REGION Network 4: Time handle
   // Es werden die Absolutwerte der Zeiten berechnet um sie dann vergleichen zu 
   // können. Intervallzeiten sind minimal 10sec. Sonst Störung "Zeitwert falsch"!
   // Bei Spaltfiltern max Laufzeit 20sec.,Min Pausenzeit 300sec.und kein Dauerbetrieb
   // möglich!
   //-----
         SET;
         R     #Temp_WrongTimevalue;
   //-----
         L     #IN_Values.RunTime;
         T     #Temp_RunTime;
         L     #IN_Values.PauseTime;
         T     #Temp_PauseTime;
   //-----
   // Absolutwerte berechnen
   //-----
         CALL  T_CONV
         ( IN  := #Temp_RunTime,
           OUT := #Temp_Runtime_ms
         );
   //-----
         CALL  T_CONV
         ( IN  := #Temp_PauseTime,
           OUT := #Temp_Pausetime_ms
         );
   //-----
         SET;
         R     #Temp_IO_Status.No_Pausetime;
   //-----
         O(;
         L     #Temp_Runtime_ms;
         L     0;
         ==I;
         );
         O(;
         L     #Temp_Pausetime_ms;
         L     0;
         ==I;
         );
         S     #Temp_IO_Status.No_Pausetime;
   //-----
   // Zeiten limitieren
   //-----
         L     #Temp_Runtime_ms;
         L     10000;  // 10 sec
         <D;
         S     #Temp_WrongTimevalue;  // Antrieb STOP!!!
         JCN   RTime;
   //-----
         L     S5T#10S;
         T     #Temp_RunTime;
   //-----
   RTime:NOP   0;
   //-----
         L     #Temp_Pausetime_ms;
         L     10000;  // 10.0 sec
         <D;
         S     #Temp_WrongTimevalue;  // Antrieb STOP!!!
   //-----
         JCN   PTime;
         L     S5T#10S;
         T     #Temp_PauseTime;
   //-----
   PTime:NOP   0;
   //-----
         O     #Temp_IO_Status.No_Pausetime;
         R     #Temp_WrongTimevalue;
   //-----
         A     #Temp_WrongTimevalue;
         AN    #Temp_IO_Fault.FLT_wrong_Timevalue;
         S     #Temp_IO_Fault.FLT_wrong_Timevalue;
         S     #IO_NewFault;
END_REGION

REGION Network 5
   //-----
         O     #Temp_IO_Fault.FLT_Motorprotection;
         O     #Temp_IO_Fault.FLT_FrequencyConverter;
         O     #Temp_IO_Fault.FLT_MaxLTripTray;
         O     #Temp_IO_Fault.FLT_wrong_Timevalue;
         =     #Temp_IO_Status.FaultLevel_3;
   //-----
END_REGION

REGION Network 6: Error handling
   //-----
         O     #Temp_IO_Fault.FLT_Motorprotection;
         O     #Temp_IO_Fault.FLT_FrequencyConverter;
         O     #Temp_IO_Fault.FLT_MaxLTripTray;
         O     #Temp_IO_Fault.FLT_wrong_Timevalue;
         O     #Temp_IO_Fault.Mes_Min_Level;
         =     #Temp_IO_Status.FLT_Exist;
   //-----
         O     #Temp_IO_Fault.FLT_Motorprotection;
         O     #Temp_IO_Fault.FLT_FrequencyConverter;
         O     #Temp_IO_Fault.FLT_MaxLTripTray;
         O     #Temp_IO_Fault.FLT_wrong_Timevalue;
         O     #Temp_IO_Fault.Mes_Min_Level;
         S     #Temp_IO_Status.Reset_Intervall;
         S     #IO_FaultLevel_3;
   //-----
END_REGION

REGION Network 7: Desicion intervall or not!
   //-----
         O(;
         A     #IN_Request_Filling;
         A     #IN_Values.Config_bit_Filling_ON;
         AN    #IN_Values.Config_bit_Filling_Int;
         );
   //-----
         O(;
         A     #IN_Request_Feed;
         A     #IN_Values.Config_bit_Charging_ON;
         AN    #IN_Values.Config_bit_Charging_Int;
         );
   //-----
         O(;
         A     #IN_Request_Cooling;
         A     #IN_Values.Config_bit_Cooling_ON;
         AN    #IN_Values.Config_bit_Cooling_Int;
         );
   //-----
         O(;
         A     #IN_Request_Heating;
         A     #IN_Values.Config_bit_Heating_ON;
         AN    #IN_Values.config_bit_Heating_Int;
         );
   //-----
         O     #Temp_IO_Status.No_Pausetime;
         S     #Temp_IO_Status.Reset_Intervall;
   //-----
END_REGION

REGION Network 8: Reset Intervall / Angefordert setzen
   //-----
         ON    #Temp_ReleaseDrive;
         ON    #IN_Release;
         O     #Temp_IO_Status.Reset_Intervall;
         R     #Temp_IO_Status.Run;
         R     #Temp_IO_Status.Pause;
         R     #Temp_IO_Status.Reset_Intervall;
   //-----
END_REGION

REGION Network 9: Wiedereinschaltsperre
   //-----
         ON    #IN_ControlVoltage;
         FP    #Temp_IO_Status.Ramp_CVoltage_Off;
         S     #Temp_IO_Status.Start_Startupdelay;
         R     #Temp_IO_Status.Disable_Start;
         R     #IN_TimerDrive;
   //-----
         ON    #IN_Values.Config_bit_Converter;
         O     #IN_TimerDrive;
         A     #Temp_IO_Status.Start_Startupdelay;
         R     #Temp_IO_Status.Disable_Start;
         R     #Temp_IO_Status.Start_Startupdelay;
   //-----
         A     #Temp_IO_Status.Start_Startupdelay;
         JCN   Lauf;
   //-----
         A     #Temp_IO_Status.Disable_Start;
         L     S5T#10S;
         SD    #IN_TimerDrive;
   //-----
         SET;
         S     #Temp_IO_Status.Disable_Start;
   //-----
         A     #IN_TimerDrive;
         A     #Temp_IO_Status.Start_Startupdelay;
         R     #Temp_IO_Status.Start_Startupdelay;
         R     #Temp_IO_Status.Disable_Start;
   //-----
END_REGION

REGION Network 10: Laufzeit
   //-----
   Lauf: NOP   0;
   //-----
         A     #Temp_ReleaseDrive;
         AN    #Temp_IO_Status.Pause;
         AN    #Temp_IO_Status.Start_Startupdelay;
         JCN   Paus;
   //-----
         A     #Temp_IO_Status.Run;
         L     #Temp_RunTime;
         SD    #IN_TimerDrive;
   //-----
         SET;
         S     #Temp_IO_Status.Run;
   //-----
         A     #IN_TimerDrive;
         JCN   Ausg;
   //-----
         SET;
         R     #Temp_IO_Status.Run;
         R     #IN_TimerDrive;
   //-----
END_REGION

REGION Network 11: Pause
   //-----
   Paus: NOP   0;
   //-----
         A     #Temp_ReleaseDrive;
         AN    #Temp_IO_Status.Run;
         AN    #Temp_IO_Status.Start_Startupdelay;
         JCN   Ausg;
   //-----
         A     #Temp_IO_Status.Pause;
         L     #Temp_PauseTime;
         SD    #IN_TimerDrive;
   //-----
         SET;
         S     #Temp_IO_Status.Pause;
   //-----
         A     #IN_TimerDrive;
         JCN   Ausg;
   //-----
         SET;
         R     #Temp_IO_Status.Pause;
         R     #IN_TimerDrive;
   //-----
END_REGION

REGION Network 12: Output mainscontactor
   //-----
   Ausg: NOP   0;
   //-----
         O(;  // generel switch ON without frequency converter
         O     #Temp_IO_Status.No_Pausetime;
         O     #Temp_IO_Status.Run;
         A     #Temp_ReleaseDrive;
         AN    #Temp_IO_Fault.Mes_Min_Level;
         AN    #Temp_IO_Fault.FLT_wrong_Timevalue;
         AN    #Temp_IO_Fault.FLT_MaxLTripTray;
         AN    #IN_Values.Config_bit_Converter;
         );
   //-----
         O(;  // generel switch ON withfrequency converter
         A     #IN_ControlVoltage;
         AN    #Temp_IO_Status.Start_Startupdelay;
         A     #IN_Values.Config_bit_Converter;
         );
         AN    #Temp_IO_Fault.FLT_Motorprotection;
   //-----
         =     #Temp_Out_MainsContactor;
         =     #OUT_MainsContactor;
   //-----
END_REGION

REGION Network 13: Ouput release frequency converter
   //-----
         O     #Temp_IO_Status.No_Pausetime;
         O     #Temp_IO_Status.Run;
         A     #Temp_ReleaseDrive;
         A     #Temp_Out_MainsContactor;
         A     #IN_Values.Config_bit_Converter;
         AN    #Temp_IO_Fault.Mes_Min_Level;
         AN    #Temp_IO_Fault.FLT_wrong_Timevalue;
         AN    #Temp_IO_Fault.FLT_MaxLTripTray;
         AN    #Temp_IO_Fault.FLT_FrequencyConverter;
         A     #IN_FaultFreqConverter;
         =     #OUT_Release_FConverter;
         =     #Temp_Release_FConverter;
   //-----
END_REGION

REGION Network 14: State of drive: 1-> ON; 2-> Faulty; 3->Selected but not ON
   //-----
         AN    #IN_Values.Config_bit_Converter;
         A     #Temp_Out_MainsContactor;
         O     #Temp_Release_FConverter;
         L     1;
         JC    tran;
   //-----
         O     #Temp_IO_Status.FLT_Exist;
         L     2;
         JC    tran;
   //-----
         AN(;
         AN    #IN_Values.Config_bit_Converter;
         A     #Temp_Out_MainsContactor;
         O     #Temp_Release_FConverter;
         );
         AN    #Temp_IO_Status.FLT_Exist;
         A     #Temp_IO_Status.Switch_Drive_ON_OFF;
         L     3;
         JC    tran;
   //-----
         L     0;
   //-----
   tran: T     #Temp_IO_Status.State_Drive;
   //-----
END_REGION

REGION Network 15: Save data
   //-----
         CALL  BLKMOV
         ( SRCBLK  := #Temp_IO_Status,
           RET_VAL := #ERROR_CODE,
           DSTBLK  := #Anyzeiger1
         );
   //-----
         CALL  BLKMOV
         ( SRCBLK  := #Temp_IO_Fault,
           RET_VAL := #ERROR_CODE,
           DSTBLK  := #Anyzeiger2
         );
   //-----
END_REGION
END_FUNCTION

FUNCTION "FC122_EdgeFilter" : Void   // FC122, STL
TITLE = Control of several auxiliary drives of a pouring machine
{ S7_Optimized_Access := 'FALSE' }
AUTHOR : KT242
FAMILY : RS_KK
NAME : Drive
VERSION : 1.5
   VAR_INPUT
      IN_Release : Bool;   // Genarelly release 0f the drive (Operation mode)
      IN_Reset_fault : Bool;   // Signal to quit fault within function block
      IN_Fault_Motorprotection : Bool;   // Input fault motorprotection of drive
      IN_DifPressure : Bool;   // Input fault difference pressure
      IN_TimerDrive : Timer;   // Timer of general timing of the drive
      Values : "UDT710_EdgeFilter";
   END_VAR
   VAR_OUTPUT
      OUT_MainsContactor : Bool;   // Ouput mainscontactor drive or frequency converter
   END_VAR
   VAR_IN_OUT
      IO_Status : ANY;   // Stores the state of the drive
      IO_NewFault : Bool;
      IO_FaultLevel_3 : Bool;
      IO_Faults : ANY;
   END_VAR
   VAR_TEMP
      Temp_IO_Status : "UDT100_EdgeFilter";
      ERROR_CODE : Int;   // Error state of systemfunction "BLKMOV" Blockmove
      Anyzeiger1 : ANY;   // Pointer to copy thr array "IO_Status" and "Temp_IO_Status"
      Anyzeiger2 : ANY;   // Pointer to copy thr array "IO_Status" and "Temp_IO_Status"
      Temp_IO_Fault : "UDT1801_EdgeFilter";
      Temp_RunTime : S5Time;   // Flag runtime drive
      Temp_PauseTime : S5Time;   // Flag pause time
      Temp_Runtime_ms : Time;   // Flag runtime drive in millisecond
      Temp_Pausetime_ms : Time;   // Flag pause time drive in millisecond
      Temp_ReleaseDrive : Bool;   // Flag release activation drive
      Temp_Fault_Drive : Bool;
      Temp_MainsContactor : Bool;
   END_VAR
BEGIN

REGION Network 1: Saved data integration
   // Änderungen:
   // -------------------------------------------------------------------------------
   // Bei der Verwendung der Umwälzpumpe als Speisepumpe wurde dieses bei Min. 
   // Füllstand ausgeshaltet, auch wenn dies im Zyklus auftrat. Hierdurch wurden dann 
   // auch die Materialpumpen abgeschaltet.
   // v.d.Geest     25.02.2003
   // -------------------------------------------------------------------------------
   // Bei einer Ansteuerung mit Frequenzumrichter wurde nicht auf die 
   // Störungsauswertung des Umrichters gewartet bevor die Freigabe gegeben wurde. 
   // Hierdurch kam es zu Störungen bei jedem einschalten des Aggregates.
   // A. Jäger      21.11.2003
   //-----
         LAR1;
         L;
         LAR2;
   //-----
         L     W[AR2, P#0.0];  // Bytes
         T     W[AR1, P#0.0];
         L     W[AR2, P#2.0];  // Amount of bytes
         T     W[AR1, P#2.0];
         L     W[AR2, P#4.0];  // Block no,
         T     W[AR1, P#4.0];
         L     D[AR2, P#6.0];  // Startadress of datas
         T     D[AR1, P#6.0];
   //-----
         CALL  BLKMOV
         ( SRCBLK  := #Anyzeiger1,
           RET_VAL := #ERROR_CODE,
           DSTBLK  := #Temp_IO_Status
         );
   //-----
         LAR1;
         L;
         LAR2;
   //-----
         L     W[AR2, P#0.0];  // Bytes
         T     W[AR1, P#0.0];
         L     W[AR2, P#2.0];  // Amount of bytes
         T     W[AR1, P#2.0];
         L     W[AR2, P#4.0];  // Block no,
         T     W[AR1, P#4.0];
         L     D[AR2, P#6.0];  // Startadress of datas
         T     D[AR1, P#6.0];
   //-----
         CALL  BLKMOV
         ( SRCBLK  := #Anyzeiger2,
           RET_VAL := #ERROR_CODE,
           DSTBLK  := #Temp_IO_Fault
         );
   //-----
END_REGION

REGION Network 2: Fault motorprotection
   //-----
         AN    #Values.Config_Exist;
         R     #Temp_IO_Fault.FLT_Motorprotection;
         R     #Temp_IO_Fault.FLT_MaxPressureDiff;
         R     #Temp_IO_Fault.FLT_wrong_Timevalue;
         R     #Temp_IO_Status.FLT_Exist;
         R     #Temp_IO_Status.Pause;
         R     #Temp_IO_Status.Run;
         JC    Ausg;
   //-----
END_REGION

REGION Network 3: Release drive
   //-----
         O     #Temp_IO_Status.Switch_Drive_ON_OFF;
         A     #IN_Release;
         =     #Temp_ReleaseDrive;
   //-----
END_REGION

REGION Network 4: Faults
   //-----
         A     #IN_Reset_fault;
         R     #Temp_IO_Fault.FLT_Motorprotection;
         R     #Temp_IO_Fault.FLT_MaxPressureDiff;
         R     #Temp_IO_Fault.FLT_wrong_Timevalue;
   //-----
         A     #IN_Fault_Motorprotection;
         AN    #Temp_IO_Fault.FLT_Motorprotection;
         S     #Temp_IO_Fault.FLT_Motorprotection;
         S     #Temp_IO_Status.Reset_Intervall;
         S     #IO_NewFault;
   //-----
         AN    #IN_DifPressure;
         A     #Values.Config_DifPress;
         A     #Temp_ReleaseDrive;
         AN    #Temp_IO_Fault.FLT_MaxPressureDiff;
         S     #Temp_IO_Fault.FLT_MaxPressureDiff;
         S     #Temp_IO_Status.Reset_Intervall;
         S     #IO_NewFault;
   //-----
END_REGION

REGION Network 5
   //-----
         O     #Temp_IO_Fault.FLT_Motorprotection;
         O     #Temp_IO_Fault.FLT_MaxPressureDiff;
         O     #Temp_IO_Fault.FLT_wrong_Timevalue;
         =     #Temp_IO_Status.FLT_Exist;
         =     #Temp_Fault_Drive;
         =     #Temp_IO_Status.FaultLevel_3;
         S     #IO_FaultLevel_3;
   //-----
END_REGION

REGION Network 6: Time handle
   // Es werden die Absolutwerte der Zeiten berechnet um sie dann vergleichen zu 
   // können. Intervallzeiten sind minimal 10sec. Sonst Störung "Zeitwert falsch"!
   // Bei Spaltfiltern max Laufzeit 20sec.,Min Pausenzeit 300sec.und kein Dauerbetrieb
   // möglich!
   //-----
         SET;
         R     #Temp_IO_Fault.FLT_wrong_Timevalue;
   //-----
         L     #Values.RunTime;
         T     #Temp_RunTime;
         L     #Values.PauseTime;
         T     #Temp_PauseTime;
   //-----
   // Absolutwerte berechnen
   //-----
         CALL  T_CONV
         ( IN  := #Temp_RunTime,
           OUT := #Temp_Runtime_ms
         );
   //-----
         CALL  T_CONV
         ( IN  := #Temp_PauseTime,
           OUT := #Temp_Pausetime_ms
         );
   //-----
   // Zeiten limitieren
   //-----
         L     #Temp_Runtime_ms;
         L     20000;  // 20.0 sec
         >D;
         S     #Temp_IO_Fault.FLT_wrong_Timevalue;  // Antrieb STOP!!!
   //-----
         JCN   RTimeS;
         L     S5T#20S;
         T     #Temp_RunTime;
   RTimeS:NOP   0;
   //-----
         L     #Temp_Pausetime_ms;
         L     L#300000;  // 300.0 sec
         <D;
         S     #Temp_IO_Fault.FLT_wrong_Timevalue;  // Antrieb STOP!!!
   //-----
         JCN   PTimeS;
         L     S5T#5M;
         T     #Temp_PauseTime;
   //-----
   PTimeS:NOP   0;
   //-----
END_REGION

REGION Network 7: Reset Intervall / Angefordert setzen
   //-----
         ON    #Temp_ReleaseDrive;
         O     #Temp_IO_Status.Reset_Intervall;
         R     #Temp_IO_Status.Run;
         R     #Temp_IO_Status.Pause;
         R     #Temp_IO_Status.Reset_Intervall;
   //-----
END_REGION

REGION Network 8: Laufzeit
   Lauf: NOP   0;
         A     #Temp_ReleaseDrive;
         AN    #Temp_IO_Status.Pause;
         JCN   Paus;
   //
         A     #Temp_IO_Status.Run;
         L     #Temp_RunTime;
         SD    #IN_TimerDrive;
   //
         SET;
         S     #Temp_IO_Status.Run;
   //
         A     #IN_TimerDrive;
         JCN   Ausg;
         SET;
         R     #Temp_IO_Status.Run;
         R     #IN_TimerDrive;
END_REGION

REGION Network 9: Pause
   Paus: NOP   0;
         A     #Temp_ReleaseDrive;
         AN    #Temp_IO_Status.Run;
         JCN   Ausg;
   //
         A     #Temp_IO_Status.Pause;
         L     #Temp_PauseTime;
         SD    #IN_TimerDrive;
   //
         SET;
         S     #Temp_IO_Status.Pause;
   //
         A     #IN_TimerDrive;
         JCN   Ausg;
         SET;
         R     #Temp_IO_Status.Pause;
         R     #IN_TimerDrive;
END_REGION

REGION Network 10: Output mainscontactor
   Ausg: NOP   0;
   //
         A     #Temp_IO_Status.Run;  // generell Eingeschaltet ohne FU
         A     #Temp_IO_Status.Switch_Drive_ON_OFF;
         A     #IN_Release;
         AN    #Temp_IO_Fault.FLT_wrong_Timevalue;
         AN    #Temp_IO_Fault.FLT_MaxPressureDiff;
         AN    #Temp_IO_Fault.FLT_Motorprotection;
         A     #Values.Config_Exist;
         =     #OUT_MainsContactor;
         =     #Temp_MainsContactor;
END_REGION

REGION Network 11: State of drive: 1-> ON; 2->Faulty; 3->Selected but not on
   //-----
         A     #Temp_MainsContactor;
         L     1;
         JC    tran;
   //-----
         A     #Temp_Fault_Drive;
         L     2;
         JC    tran;
   //-----
         A     #Temp_IO_Status.Switch_Drive_ON_OFF;
         L     3;
         JC    tran;
   //-----
         L     0;
   //-----
   tran: T     #Temp_IO_Status.State_Drive;
END_REGION

REGION Network 12: Save data
         CALL  BLKMOV
         ( SRCBLK  := #Temp_IO_Status,
           RET_VAL := #ERROR_CODE,
           DSTBLK  := #Anyzeiger1
         );
   //
         CALL  BLKMOV
         ( SRCBLK  := #Temp_IO_Fault,
           RET_VAL := #ERROR_CODE,
           DSTBLK  := #Anyzeiger2
         );
   //
END_REGION
END_FUNCTION

FUNCTION "FC123_FeedingPump" : Void   // FC123, STL
TITLE = Control of several auxiliary drives of a pouring machine
{ S7_Optimized_Access := 'FALSE' }
AUTHOR : KT242
FAMILY : RS_KK
NAME : Drive
VERSION : 1.5
   VAR_INPUT
      IN_Release : Bool;   // Genarelly release 0f the drive (Operation mode)
      IN_ControlVoltage : Bool;   // Signal delay activation frequency converter (protection after emergency-stop)
      IN_Reset_fault : Bool;   // Signal to quit fault within function block
      IN_ComponentDeselected : Bool;   // is the component deselected? -> Fault Group 1 -> Groupe 3
      IN_Request_Feed : Bool;   // Request switch on drive if componenten pump start up
      IN_Request_Filling : Bool;   // Request switch on drive for filling
      IN_Request_Bypass : Bool;   // Request switch on drive for bypass circulation
      IN_Fault_Motorprotection : Bool;   // Input fault motorprotection of drive
      IN_FaultFreqConverter : Bool;   // Input fault frequency converter of drive
      IN_DryRun : Bool;   // Input fault Min_Level or dry run
      IN_MaxLevelTray : Bool;   // Input fault max. filling level tray
      IN_MaxPressure : Bool;   // Input Max pressure switch
      IN_TempRelease : Bool;   // Input Min. Temperature reacht for switch on
      IN_TimerDrive : Timer;   // Timer of general timing of the drive
      IN_TimerStartUpFConv : Timer;   // Timer of delay start up frequency converter
      Values : "UDT710_FeedingPump";
   END_VAR
   VAR_OUTPUT
      OUT_MainsContactor : Bool;   // Ouput mainscontactor drive or frequency converter
      OUT_Release_FConverter : Bool;   // Output release of frequncy converter to control rotation speed
   END_VAR
   VAR_IN_OUT
      IO_Status : ANY;   // Stores the state of the drive
      IO_NewFault : Bool;
      IO_FaultLevel_1 : Bool;
      IO_FaultLevel_3 : Bool;
      IO_Faults : ANY;
   END_VAR
   VAR_TEMP
      Temp_IO_Status : "UDT100_FeedingPump";
      ERROR_CODE : Int;   // Error state of systemfunction "BLKMOV" Blockmove
      Anyzeiger1 : ANY;   // Pointer to copy thr array "IO_Status" and "Temp_IO_Status"
      Anyzeiger2 : ANY;   // Pointer to copy thr array "IO_Status" and "Temp_IO_Status"
      Temp_IO_Fault : "UDT1801_FeedingPump";
      Temp_RunTime : S5Time;   // Flag runtime drive
      Temp_PauseTime : S5Time;   // Flag pause time
      Temp_Runtime_ms : Time;   // Flag runtime drive in millisecond
      Temp_Pausetime_ms : Time;   // Flag pause time drive in millisecond
      Temp_ReleaseDrive : Bool;   // Flag release activation drive
      Temp_Fault_Drive : Bool;
      Temp_WrongTimevalue : Bool;
      Temp_MainsContactor : Bool;
      Temp_Release_FConverter : Bool;
   END_VAR
BEGIN

REGION Network 1: Saved data integration
   // Änderungen:
   // -------------------------------------------------------------------------------
   // Bei der Verwendung der Umwälzpumpe als Speisepumpe wurde dieses bei Min. 
   // Füllstand ausgeshaltet, auch wenn dies im Zyklus auftrat. Hierdurch wurden dann 
   // auch die Materialpumpen abgeschaltet.
   // v.d.Geest     25.02.2003
   // -------------------------------------------------------------------------------
   // Bei einer Ansteuerung mit Frequenzumrichter wurde nicht auf die 
   // Störungsauswertung des Umrichters gewartet bevor die Freigabe gegeben wurde. 
   // Hierdurch kam es zu Störungen bei jedem einschalten des Aggregates.
   // A. Jäger      21.11.2003
   //-----
         LAR1;
         L;
         LAR2;
   //-----
         L     W[AR2, P#0.0];  // Bytes
         T     W[AR1, P#0.0];
         L     W[AR2, P#2.0];  // Amount of bytes
         T     W[AR1, P#2.0];
         L     W[AR2, P#4.0];  // Block no,
         T     W[AR1, P#4.0];
         L     D[AR2, P#6.0];  // Startadress of datas
         T     D[AR1, P#6.0];
   //-----
         CALL  BLKMOV
         ( SRCBLK  := #Anyzeiger1,
           RET_VAL := #ERROR_CODE,
           DSTBLK  := #Temp_IO_Status
         );
   //-----
         LAR1;
         L;
         LAR2;
   //-----
         L     W[AR2, P#0.0];  // Bytes
         T     W[AR1, P#0.0];
         L     W[AR2, P#2.0];  // Amount of bytes
         T     W[AR1, P#2.0];
         L     W[AR2, P#4.0];  // Block no,
         T     W[AR1, P#4.0];
         L     D[AR2, P#6.0];  // Startadress of datas
         T     D[AR1, P#6.0];
   //-----
         CALL  BLKMOV
         ( SRCBLK  := #Anyzeiger2,
           RET_VAL := #ERROR_CODE,
           DSTBLK  := #Temp_IO_Fault
         );
   //-----
END_REGION

REGION Network 2: Fault motorprotection
   //-----
         AN    #Values.Config_Exist;
         R     #Temp_IO_Fault.FLT_Motorprotection;
         R     #Temp_IO_Fault.FLT_FrequencyConverter;
         R     #Temp_IO_Fault.FLT_MaxLTripTray;
         R     #Temp_IO_Fault.FLT_Dryrunsafety;
         R     #Temp_IO_Fault.FLT_wrong_Timevalue;
         R     #Temp_IO_Fault.FLT_MaxPressure;
         R     #Temp_IO_Fault.Mes_Min_temp;
         R     #Temp_IO_Status.FLT_Exist;
         R     #Temp_IO_Status.Pause;
         R     #Temp_IO_Status.Run;
         JC    Ausg;
   //-----
END_REGION

REGION Network 3: Release drive
   //-----
         O(;
         A     #IN_Request_Filling;
         A     #Values.Config_Filling;
         A     #Temp_IO_Status.Switch_Drive_ON_OFF;
         );
         O(;
         A     #IN_Request_Bypass;
         A     #Values.Config_Bypass;
         A     #Temp_IO_Status.Switch_Drive_ON_OFF;
         );
         O(;
         A     #Temp_IO_Status.Switch_Drive_ON_OFF;
         A     #Values.Config_ManualSwitchON;
         );
         O(;
         A     #IN_Request_Feed;
         );
         A     #IN_Release;
         =     #Temp_ReleaseDrive;
   //-----
END_REGION

REGION Network 4: Faults
   //-----
         A     #IN_Reset_fault;
         R     #Temp_IO_Fault.FLT_Motorprotection;
         R     #Temp_IO_Fault.FLT_FrequencyConverter;
         R     #Temp_IO_Fault.FLT_MaxLTripTray;
         R     #Temp_IO_Fault.FLT_Dryrunsafety;
         R     #Temp_IO_Fault.FLT_wrong_Timevalue;
         R     #Temp_IO_Fault.FLT_MaxPressure;
   //-----
         A     #IN_Fault_Motorprotection;
         AN    #Temp_IO_Fault.FLT_Motorprotection;
         S     #Temp_IO_Fault.FLT_Motorprotection;
         S     #IO_NewFault;
   //-----
         A     #IN_ControlVoltage;
         AN    #Temp_IO_Fault.FLT_wrong_Timevalue;
         AN    #Temp_IO_Status.Start_Startupdelay;
         L     S5T#5S;
         SD    #IN_TimerStartUpFConv;
   //-----
         A     #IN_TimerStartUpFConv;
         AN    #IN_FaultFreqConverter;
         A     #Temp_ReleaseDrive;
         A     #Values.Config_WithFC;
         AN    #Temp_IO_Fault.FLT_FrequencyConverter;
         S     #Temp_IO_Fault.FLT_FrequencyConverter;
         S     #IO_NewFault;
   //-----
         AN    #IN_MaxLevelTray;
         A     #Temp_ReleaseDrive;
         AN    #Temp_IO_Fault.FLT_MaxLTripTray;
         S     #Temp_IO_Fault.FLT_MaxLTripTray;
         S     #IO_NewFault;
   //-----
         AN    #IN_DryRun;
         A     #Temp_ReleaseDrive;
         AN    #Temp_IO_Fault.FLT_Dryrunsafety;
         S     #Temp_IO_Fault.FLT_Dryrunsafety;
         S     #IO_NewFault;
   //-----
         AN    #IN_MaxPressure;
         AN    #Temp_IO_Fault.FLT_MaxPressure;
         S     #Temp_IO_Fault.FLT_MaxPressure;
         S     #IO_NewFault;
   //-----
         AN    #IN_TempRelease;
         A     #Temp_ReleaseDrive;
         AN    #Temp_IO_Fault.Mes_Min_temp;
         S     #Temp_IO_Fault.Mes_Min_temp;
         S     #IO_NewFault;
   //-----
         A     #IN_TempRelease;
         ON    #Temp_ReleaseDrive;
         R     #Temp_IO_Fault.Mes_Min_temp;
   //-----
         A     #Temp_IO_Fault.Mes_Min_temp;
         R     #Temp_ReleaseDrive;
   //-----
END_REGION

REGION Network 5: A fault group 1 exist
   //-----
         O     #Temp_IO_Fault.FLT_MaxLTripTray;
         O     #Temp_IO_Fault.FLT_MaxPressure;
         O     #Temp_IO_Fault.FLT_Dryrunsafety;
         AN    #IN_ComponentDeselected;
         =     #Temp_IO_Status.FaultLevel_1;
   //-----
         O     #Temp_IO_Fault.FLT_MaxLTripTray;
         O     #Temp_IO_Fault.FLT_MaxPressure;
         O     #Temp_IO_Fault.FLT_Dryrunsafety;
         A     #IN_ComponentDeselected;
         O     #Temp_IO_Fault.FLT_Motorprotection;
         O     #Temp_IO_Fault.FLT_FrequencyConverter;
         O     #Temp_IO_Fault.FLT_wrong_Timevalue;
         =     #Temp_IO_Status.FaultLevel_3;
   //-----
END_REGION

REGION Network 6: Time handle
   // Es werden die Absolutwerte der Zeiten berechnet um sie dann vergleichen zu 
   // können. Intervallzeiten sind minimal 10sec. Sonst Störung "Zeitwert falsch"!
   // Bei Spaltfiltern max Laufzeit 20sec.,Min Pausenzeit 300sec.und kein Dauerbetrieb
   // möglich!
   //-----
         SET;
         R     #Temp_WrongTimevalue;
   //-----
         L     #Values.RunTime;
         T     #Temp_RunTime;
         L     #Values.PauseTime;
         T     #Temp_PauseTime;
   //-----
   // Absolutwerte berechnen
   //-----
         CALL  T_CONV
         ( IN  := #Temp_RunTime,
           OUT := #Temp_Runtime_ms
         );
   //-----
         CALL  T_CONV
         ( IN  := #Temp_PauseTime,
           OUT := #Temp_Pausetime_ms
         );
   //-----
         SET;
         R     #Temp_IO_Status.No_Pausetime;
   //-----
         O(;
         L     #Temp_Runtime_ms;
         L     0;
         ==I;
         );
         O(;
         L     #Temp_Pausetime_ms;
         L     0;
         ==I;
         );
         S     #Temp_IO_Status.No_Pausetime;
   //-----
   // Zeiten limitieren
   //-----
         L     #Temp_Runtime_ms;
         L     10000;  // 10 sec
         <D;
         S     #Temp_WrongTimevalue;  // Antrieb STOP!!!
         JCN   nLi1;
   //-----
         L     S5T#10S;
         T     #Temp_RunTime;
   //-----
   nLi1: L     #Temp_Pausetime_ms;
         L     10000;  // 10.0 sec
         <D;
         S     #Temp_WrongTimevalue;  // Antrieb STOP!!!
         JCN   nLi2;
   //-----
         L     S5T#10S;
         T     #Temp_PauseTime;
         JU    nLi2;
   //-----
   nLi2: NOP   0;
   //-----
         AN    #Temp_WrongTimevalue;
         R     #Temp_IO_Fault.FLT_wrong_Timevalue;
   //-----
         A     #Temp_WrongTimevalue;
         AN    #Temp_IO_Status.No_Pausetime;
         AN    #Temp_IO_Fault.FLT_wrong_Timevalue;
         S     #Temp_IO_Fault.FLT_wrong_Timevalue;
         S     #IO_NewFault;
   //-----
END_REGION

REGION Network 7: Error handling
   //-----
         O     #Temp_IO_Fault.FLT_Motorprotection;
         O     #Temp_IO_Fault.FLT_FrequencyConverter;
         O     #Temp_IO_Fault.FLT_MaxLTripTray;
         O     #Temp_IO_Fault.FLT_Dryrunsafety;
         O     #Temp_IO_Fault.FLT_wrong_Timevalue;
         =     #Temp_IO_Status.FLT_Exist;
         =     #Temp_Fault_Drive;
   //-----
         O     #Temp_IO_Fault.FLT_Motorprotection;
         O     #Temp_IO_Fault.FLT_FrequencyConverter;
         O     #Temp_IO_Fault.FLT_Dryrunsafety;
         O     #Temp_IO_Fault.FLT_MaxLTripTray;
         O     #Temp_IO_Fault.FLT_wrong_Timevalue;
         S     #Temp_IO_Status.Reset_Intervall;
         S     #IO_FaultLevel_3;
   //-----
END_REGION

REGION Network 8: Desicion intervall or not!
         O(;
         A     #IN_Request_Filling;
         A     #Values.Config_Filling;
         A     #Temp_IO_Status.Switch_Drive_ON_OFF;
         );
         O     #IN_Request_Feed;
         O     #Temp_IO_Status.No_Pausetime;
         S     #Temp_IO_Status.Reset_Intervall;
END_REGION

REGION Network 9: Reset Intervall / Angefordert setzen
   //-----
         ON    #Temp_ReleaseDrive;
         ON    #IN_Release;
         O     #Temp_IO_Status.Reset_Intervall;
         R     #Temp_IO_Status.Run;
         R     #Temp_IO_Status.Pause;
         R     #Temp_IO_Status.Reset_Intervall;
   //-----
END_REGION

REGION Network 10: Wiedereinschaltsperre
   //-----
         ON    #IN_ControlVoltage;
         FP    #Temp_IO_Status.Ramp_CVoltage_Off;
         S     #Temp_IO_Status.Start_Startupdelay;
         R     #Temp_IO_Status.Disable_Start;
         R     #IN_TimerDrive;
   //-----
         ON    #Values.Config_WithFC;
         O     #IN_TimerDrive;
         A     #Temp_IO_Status.Start_Startupdelay;
         R     #Temp_IO_Status.Disable_Start;
         R     #Temp_IO_Status.Start_Startupdelay;
   //-----
         A     #Temp_IO_Status.Start_Startupdelay;
         JCN   Lauf;
   //-----
         A     #Temp_IO_Status.Disable_Start;
         L     S5T#10S;
         SD    #IN_TimerDrive;
   //-----
         SET;
         S     #Temp_IO_Status.Disable_Start;
   //-----
         A     #IN_TimerDrive;
         A     #Temp_IO_Status.Start_Startupdelay;
         R     #Temp_IO_Status.Start_Startupdelay;
         R     #Temp_IO_Status.Disable_Start;
   //-----
END_REGION

REGION Network 11: Laufzeit
   Lauf: NOP   0;
         A     #Temp_ReleaseDrive;
         AN    #Temp_IO_Status.Pause;
         AN    #Temp_IO_Status.Start_Startupdelay;
         JCN   Paus;
   //
         A     #Temp_IO_Status.Run;
         L     #Temp_RunTime;
         SD    #IN_TimerDrive;
   //
         SET;
         S     #Temp_IO_Status.Run;
   //
         A     #IN_TimerDrive;
         JCN   Ausg;
         SET;
         R     #Temp_IO_Status.Run;
         R     #IN_TimerDrive;
END_REGION

REGION Network 12: Pause
   //-----
   Paus: NOP   0;
   //-----
         A     #Temp_ReleaseDrive;
         AN    #Temp_IO_Status.Run;
         AN    #Temp_IO_Status.Start_Startupdelay;
         JCN   Ausg;
   //-----
         A     #Temp_IO_Status.Pause;
         L     #Temp_PauseTime;
         SD    #IN_TimerDrive;
   //-----
         SET;
         S     #Temp_IO_Status.Pause;
   //-----
         A     #IN_TimerDrive;
         JCN   Ausg;
   //-----
         SET;
         R     #Temp_IO_Status.Pause;
         R     #IN_TimerDrive;
   //-----
END_REGION

REGION Network 13: Output mainscontactor
   //-----
   Ausg: NOP   0;
   //-----
         O(;  // generel switch ON without frequency converter
         O     #Temp_IO_Status.No_Pausetime;
         O     #Temp_IO_Status.Run;
         A     #Temp_ReleaseDrive;
         A(;  // If Filling is aktiv the dryrun must switched
         A     #IN_Request_Filling;
         A     #Values.Config_Filling;
         A     #Temp_IO_Status.Switch_Drive_ON_OFF;
         ON    #Temp_IO_Fault.FLT_Dryrunsafety;
         );
         AN    #Temp_IO_Fault.FLT_wrong_Timevalue;
         AN    #Temp_IO_Fault.FLT_MaxLTripTray;
         AN    #Values.Config_WithFC;
         );
         O(;  // generel switch ON withfrequency converter
         A     #IN_ControlVoltage;
         AN    #Temp_IO_Status.Start_Startupdelay;
         A     #Values.Config_WithFC;
         );
         AN    #Temp_IO_Fault.FLT_Motorprotection;
         A     #Values.Config_Exist;
   //-----
         =     #OUT_MainsContactor;
         =     #Temp_MainsContactor;
   //-----
END_REGION

REGION Network 14: Ouput release frequency converter
   //-----
         O     #Temp_IO_Status.No_Pausetime;
         O     #Temp_IO_Status.Run;
         A     #Temp_ReleaseDrive;
         A     #Temp_MainsContactor;
         A     #Values.Config_WithFC;
         A(;  // If Filling is aktiv the dryrun must switched
         A     #IN_Request_Filling;
         A     #Values.Config_Filling;
         A     #Temp_IO_Status.Switch_Drive_ON_OFF;
         ON    #Temp_IO_Fault.FLT_Dryrunsafety;
         );
         AN    #Temp_IO_Fault.FLT_wrong_Timevalue;
         AN    #Temp_IO_Fault.FLT_MaxLTripTray;
         AN    #Temp_IO_Fault.FLT_FrequencyConverter;
         A     #IN_FaultFreqConverter;
         A     #Values.Config_Exist;
         =     #OUT_Release_FConverter;
         =     #Temp_Release_FConverter;
   //-----
END_REGION

REGION Network 15: State of drive: 1-> ON; 2-> Faulty; 3->Selected but not ON
   //-----
         AN    #Values.Config_WithFC;
         A     #Temp_MainsContactor;
         O     #Temp_Release_FConverter;
         L     1;
         JC    tran;
   //-----
         A     #Temp_Fault_Drive;
         L     2;
         JC    tran;
   //-----
         A     #Temp_IO_Status.Switch_Drive_ON_OFF;
         L     3;
         JC    tran;
   //-----
         L     0;
   //-----
   tran: T     #Temp_IO_Status.State_Drive;
   //-----
END_REGION

REGION Network 16: Save data
   //-----
         CALL  BLKMOV
         ( SRCBLK  := #Temp_IO_Status,
           RET_VAL := #ERROR_CODE,
           DSTBLK  := #Anyzeiger1
         );
   //-----
         CALL  BLKMOV
         ( SRCBLK  := #Temp_IO_Fault,
           RET_VAL := #ERROR_CODE,
           DSTBLK  := #Anyzeiger2
         );
   //-----
END_REGION
END_FUNCTION

FUNCTION "FC126_write_ProCan" : Void   // FC126, STL
TITLE = Write to IO-Interface of ProCan modul
{ S7_Optimized_Access := 'FALSE' }
AUTHOR : KT242
FAMILY : RS_KK
NAME : WRProcan
VERSION : 1.1
   VAR_TEMP
      Nullmerker : Byte;   // Zwischenmerker mit dem Wert "0" zum ablöschen bei gestörter Übertragung
      ERROR_CODE : DInt;   // Störungszustand der Systemfunktion "FILL" Blockmove
      Temp_ToolAdr : Int;
      Temp_PS_offset : Int;
      TempShotWithMaterial_M1 : Bool;
      TempShotWithMaterial_M2 : Bool;
      Temp_OperationMode : Bool;
      ControlBitShot : Byte;
      Temp_MH_OutputSignals : Word;
      TempMH_Bit : DWord;
      Temp_MH_Shot_MH01 : Bool;
      Temp_MH_Shot_MH02 : Bool;
      Temp_MH_Shot_MH03 : Bool;
      Temp_MH_Shot_MH04 : Bool;
      Temp_MH_Shot_MH05 : Bool;
      Temp_MH_Shot_MH06 : Bool;
      Temp_MH_Shot_MH07 : Bool;
      Temp_MH_Shot_MH08 : Bool;
      Temp_MH_Shot_MH09 : Bool;
      Temp_MH_Shot_MH10 : Bool;
      Temp_CorrValue : Real;
      Temp_Error : Bool;
      TempFlowIndex : Byte;
      TemRetBLKMOV : Int;
      TempTandem : Word;
      Dummy : Bool;
      TempNozzelBitCirc : Byte;
      TempNozzelBitShot : Byte;
      TempAdrNozzel : Int;
      TempNozzelBitForce : Byte;
      ControlByteCtrlCP : Byte;
      ThrottleGap : Int;
      TempNozzelBitRelease : Byte;
      ShotTime_M1 : DInt;
      ControlFlowIndex : Byte;
      ControlBitCP : Byte;
      Temp_CycleRunning : Array[1..16] of Bool;
   END_VAR
BEGIN

REGION Network 1: Write data flow 1
   //----------------------------------------------------------------------
   // Check if the communication partner is ready for
   // data transfer to ProCan
   // ---------------------------------------------------------------------
         AN    "PN_FlowRate".Component[1].FlowC_F.Active;
         JC    ed01;
   //-----------------------------------------------------------------
   // Flow set value
   //-----------------------------------------------------------------
         L     0;
         L     "PN_FlowRate".Component[1].FlowC_F.Address;
         <>D;
         JCN   qp01;
         SLD   3;
         LAR1;
         L     0;
         A     "TM_pulse_2PointAdjust_C1";
         JC    _2point_C1;
         L     "DB613_Komponent_State".FlowPump[1];
   _2point_C1:T     PQD [ AR1 , P#0.0 ];

   //---------------------------------------------------------------------
   // Quick pressure build up
   //---------------------------------------------------------------------
   qp01: L     0;
         L     "PN_FlowRate".Component[1].FlowC_F.Address;
         <>D;
         JCN   fi01;
         L     4;
         +D;
         SLD   3;
         LAR1;
         L     "DB613_Komponent_State".FlowPumpQPB[1];
         T     PQD[AR1, P#0.0];

         L     0;
         L     "PN_FlowRate".Component[1].FlowC_F.Address;
         <>D;
         JCN   fi01;
         L     8;
         +D;
         SLD   3;
         LAR1;
         L     "DB613_Komponent_State".PressurePumpQPB[1];
         T     PQD [ AR1 , P#0.0 ];

   //--- Pressure from external device ???
   //    L     0
   //    L     "DB1233_ProCanIO_Flow".AddressFlow[1].Ref_Act_PressureQPB
   //    <I
   //    SPBN  fi01
   //    SLD   3
   //    LAR1
   //    L     DB60.DBW    2
   //    L     10
   //    *D
   //    T     PAW [AR1,P#0.0]

   //-----------------------------------------------------------------
   // Flow-Index: Enableclosedloop; Start quick pressure build up
   //-----------------------------------------------------------------
   fi01: L     0;
         T     #ControlFlowIndex;

   //-----------------------------------------
   // Enableclosedloop
   //-----------------------------------------
         AN    "DB613_Komponent_State".MeteringPump[1].Enableclosedloop;
         JC    SDA1;
         L     2#0000_0010;
         L     #ControlFlowIndex;
         OW;
         T     #ControlFlowIndex;

   //-----------------------------------------
   // Trigger SDA
   //-----------------------------------------
   SDA1: ON    "DB613_Komponent_State".MeteringPump[1].Puls_SDA;
         O(;
         L     "DB613_Komponent_State".FlowPumpQPB[1];
         L     0.0;
         ==R;
         );
         O(;
         L     "DB613_Komponent_State".PressurePumpQPB[1];
         L     0.0;
         ==R;
         );
         JC    TAB1;
         L     2#0000_1000;
         L     #ControlFlowIndex;
         OW;
         T     #ControlFlowIndex;

   //-----------------------------------------
   // Write Output
   //-----------------------------------------
   TAB1: L     0;
         L     "PN_FlowRate".Component[1].FlowC_F.Address;
         <>D;
         JCN   ed01;
         L     16;
         +D;
         SLD   3;
         LAR1;
         L     #ControlFlowIndex;
         T     PQB [ AR1 , P#0.0 ];

   //----------------------------------------------------------------
   // Tandem comand
   //----------------------------------------------------------------
   ta01: NOP   0;
   //      L     0
   //      L     "DB1233_ProCanIO_Flow".AddressFlow[1].Ref_TandemComand
   //      <I
   //      SPBN  ed01
   //      SLD   3
   //      LAR1
   //
   //      CALL  BLKMOV
   //         blk_type:=Any
   //         SRCBLK  :="DB206_TandemCommand".PistonPair[1]
   //         RET_VAL :=#TemRetBLKMOV
   //         DSTBLK  :=#TempTandem
   //
   //      L     #TempTandem
   //      TAW
   //      T PAB [ AR1 , P#0.0 ]

   ed01: NOP   0;
END_REGION

REGION Network 2: Write data flow 2
   //----------------------------------------------------------------------
   // Check if the communication partner is ready for
   // data transfer to ProNet
   // ---------------------------------------------------------------------
         AN    "PN_FlowRate".Component[2].FlowC_F.Active;
         JC    ed02;
   //-----------------------------------------------------------------
   // Flow set value
   //-----------------------------------------------------------------
         L     0;
         L     "PN_FlowRate".Component[2].FlowC_F.Address;
         <>D;
         JCN   qp02;
         SLD   3;
         LAR1;
         L     0;
         A     "TM_pulse_2PointAdjust_C2";
         JC    _2point_C2;
         L     "DB613_Komponent_State".FlowPump[2];
   _2point_C2:T     PQD [ AR1 , P#0.0 ];


   //---------------------------------------------------------------------
   // Quick pressure build up
   //---------------------------------------------------------------------
   qp02: L     0;
         L     "PN_FlowRate".Component[2].FlowC_F.Address;
         <>D;
         JCN   fi02;
         L     4;
         +D;
         SLD   3;
         LAR1;
         L     "DB613_Komponent_State".FlowPumpQPB[2];
         T     PQD[AR1, P#0.0];

         L     0;
         L     "PN_FlowRate".Component[2].FlowC_F.Address;
         <>D;
         JCN   fi02;
         L     8;
         +D;
         SLD   3;
         LAR1;
         L     "DB613_Komponent_State".PressurePumpQPB[2];
         T     PQD [ AR1 , P#0.0 ];

   //--- Pressure from external device ???
   //    L     0
   //    L     "DB1233_ProCanIO_Flow".AddressFlow[2].Ref_Act_PressureQPB
   //    <I
   //    SPBN  fi01
   //    SLD   3
   //    LAR1
   //    L     DB60.DBW    2
   //    L     10
   //    *D
   //    T     PAW [AR1,P#0.0]

   //-----------------------------------------------------------------
   // Flow-Index: Enableclosedloop; Start quick pressure build up
   //-----------------------------------------------------------------
   fi02: L     0;
         T     #ControlFlowIndex;

   //-----------------------------------------
   // Enableclosedloop
   //-----------------------------------------
         AN    "DB613_Komponent_State".MeteringPump[2].Enableclosedloop;
         JC    SDA2;
         L     2#0000_0010;
         L     #ControlFlowIndex;
         OW;
         T     #ControlFlowIndex;

   //-----------------------------------------
   // Trigger SDA
   //-----------------------------------------
   SDA2: ON    "DB613_Komponent_State".MeteringPump[2].Puls_SDA;
         O(;
         L     "DB613_Komponent_State".FlowPumpQPB[2];
         L     0.0;
         ==R;
         );
         O(;
         L     "DB613_Komponent_State".PressurePumpQPB[2];
         L     0.0;
         ==R;
         );
         JC    TAB2;
         L     2#0000_1000;
         L     #ControlFlowIndex;
         OW;
         T     #ControlFlowIndex;

   //-----------------------------------------
   // Write Output
   //-----------------------------------------
   TAB2: L     0;
         L     "PN_FlowRate".Component[2].FlowC_F.Address;
         <>D;
         JCN   ed02;
         L     16;
         +D;
         SLD   3;
         LAR1;
         L     #ControlFlowIndex;
         T     PQB [ AR1 , P#0.0 ];

   //----------------------------------------------------------------
   // Tandem comand
   //----------------------------------------------------------------
   ta02: NOP   0;
   //      L     0
   //      L     "DB1233_ProCanIO_Flow".AddressFlow[2].Ref_TandemComand
   //      <I
   //      SPBN  ed02
   //      SLD   3
   //      LAR1
   //
   //      CALL  BLKMOV
   //         blk_type:=Any
   //         SRCBLK  :="DB206_TandemCommand".PistonPair[2]
   //         RET_VAL :=#TemRetBLKMOV
   //         DSTBLK  :=#TempTandem
   //
   //      L     #TempTandem
   //      TAW
   //      T PAB [ AR1 , P#0.0 ]

   ed02: NOP   0;
END_REGION

REGION Network 3: Write data flow 3
   //----------------------------------------------------------------------
   // Check if the communication partner is ready for
   // data transfer to ProNet
   // ---------------------------------------------------------------------
         AN    "PN_FlowRate".Component[3].FlowC_F.Active;
         JC    ed03;
   //-----------------------------------------------------------------
   // Flow set value
   //-----------------------------------------------------------------
         L     0;
         L     "PN_FlowRate".Component[3].FlowC_F.Address;
         <>D;
         JCN   qp03;
         SLD   3;
         LAR1;
         L     "DB613_Komponent_State".FlowPump[3];
         T     PQD[AR1, P#0.0];

   //---------------------------------------------------------------------
   // Quick pressure build up
   //---------------------------------------------------------------------
   qp03: L     0;
         L     "PN_FlowRate".Component[3].FlowC_F.Address;
         <>D;
         JCN   fi03;
         L     4;
         +D;
         SLD   3;
         LAR1;
         L     "DB613_Komponent_State".FlowPumpQPB[3];
         T     PQD[AR1, P#0.0];

         L     0;
         L     "PN_FlowRate".Component[3].FlowC_F.Address;
         <>D;
         JCN   fi03;
         L     8;
         +D;
         SLD   3;
         LAR1;
         L     "DB613_Komponent_State".PressurePumpQPB[3];
         T     PQD [ AR1 , P#0.0 ];

   //--- Pressure from external device ???
   //    L     0
   //    L     "DB1233_ProCanIO_Flow".AddressFlow[3].Ref_Act_PressureQPB
   //    <I
   //    SPBN  fi01
   //    SLD   3
   //    LAR1
   //    L     DB60.DBW    2
   //    L     10
   //    *D
   //    T     PAW [AR1,P#0.0]

   //-----------------------------------------------------------------
   // Flow-Index: Enableclosedloop; Start quick pressure build up
   //-----------------------------------------------------------------
   fi03: L     0;
         T     #ControlFlowIndex;

   //-----------------------------------------
   // Enableclosedloop
   //-----------------------------------------
         AN    "DB613_Komponent_State".MeteringPump[3].Enableclosedloop;
         JC    SDA3;
         L     2#0000_0010;
         L     #ControlFlowIndex;
         OW;
         T     #ControlFlowIndex;

   //-----------------------------------------
   // Trigger SDA
   //-----------------------------------------
   SDA3: ON    "DB613_Komponent_State".MeteringPump[3].Puls_SDA;
         O(;
         L     "DB613_Komponent_State".FlowPumpQPB[3];
         L     0.0;
         ==R;
         );
         O(;
         L     "DB613_Komponent_State".PressurePumpQPB[3];
         L     0.0;
         ==R;
         );
         JC    TAB3;
         L     2#0000_1000;
         L     #ControlFlowIndex;
         OW;
         T     #ControlFlowIndex;

   //-----------------------------------------
   // Write Output
   //-----------------------------------------
   TAB3: L     0;
         L     "PN_FlowRate".Component[3].FlowC_F.Address;
         <>D;
         JCN   ed03;
         L     16;
         +D;
         SLD   3;
         LAR1;
         L     #ControlFlowIndex;
         T     PQB [ AR1 , P#0.0 ];

   //----------------------------------------------------------------
   // Tandem comand  (DB206 has to be expanded)
   //----------------------------------------------------------------
   ta03: NOP   0;
   //      L     0
   //      L     "DB1233_ProCanIO_Flow".AddressFlow[3].Ref_TandemComand
   //      <I
   //      SPBN  ed03
   //      SLD   3
   //      LAR1

   //      CALL  "BLKMOV"
   //       SRCBLK :="DB206_TandemCommand"
   //       RET_VAL:=#TemRetBLKMOV
   //       DSTBLK :=#TempTandem

   //      L     #TempTandem
   //      TAW
   //      T     PAB [AR1,P#0.0]
   ed03: NOP   0;
END_REGION

REGION Network 4: Write data flow 4
   //----------------------------------------------------------------------
   // Check if the communication partner is ready for
   // data transfer to ProCan
   // ---------------------------------------------------------------------
         AN    "PN_FlowRate".Component[4].FlowC_F.Active;
         JC    ed04;
   //-----------------------------------------------------------------
   // Flow set value
   //-----------------------------------------------------------------
         L     0;
         L     "PN_FlowRate".Component[4].FlowC_F.Address;
         <>D;
         JCN   qp04;
         SLD   3;
         LAR1;
         L     "DB613_Komponent_State".FlowPump[4];
         T     PQD[AR1, P#0.0];

   //---------------------------------------------------------------------
   // Quick pressure build up
   //---------------------------------------------------------------------
   qp04: L     0;
         L     "PN_FlowRate".Component[4].FlowC_F.Address;
         <>D;
         JCN   fi04;
         L     4;
         +D;
         SLD   3;
         LAR1;
         L     "DB613_Komponent_State".FlowPumpQPB[4];
         T     PQD[AR1, P#0.0];

         L     0;
         L     "PN_FlowRate".Component[4].FlowC_F.Address;
         <>D;
         JCN   fi04;
         L     8;
         +D;
         SLD   3;
         LAR1;
         L     "DB613_Komponent_State".PressurePumpQPB[4];
         T     PQW[AR1, P#0.0];

   //--- Pressure from external device ???
   //    L     0
   //    L     "DB1233_ProCanIO_Flow".AddressFlow[4].Ref_Act_PressureQPB
   //    <I
   //    SPBN  fi04
   //    SLD   3
   //    LAR1
   //    L     DB60.DBW    2
   //    L     10
   //    *D
   //    T     PAW [AR1,P#0.0]

   //-----------------------------------------------------------------
   // Flow-Index: Enableclosedloop; Start quick pressure build up
   //-----------------------------------------------------------------
   fi04: L     0;
         T     #ControlFlowIndex;